// Mitsubishi GX Works2 project: 70常温静置库1130   PLC: Q10UDEH

TYPE BatteryCode : STRUCT
  arrwCode : ARRAY [0..8] OF WORD;
END_STRUCT END_TYPE

TYPE CommunicationIO : STRUCT
  i_iResponsPCPLC : INT;  (* 上位机写入-请求确认 *)
  i_iReadWriteFlagPCPLC : INT;  (* 上位机写入-读写标志位 *)
  i_iTaskProcessFlagPCPLC : INT;  (* 上位机写入-任务处理标志位 *)
  i_iCommandPCPLC : INT;  (* 上位机写入-命令字 *)
  i_iTaskIDPCPLC : INT;  (* 上位机写入-任务号 *)
  i_diDestinationDevicePCPLC : DINT;  (* 上位机写入-目标设备号 *)
  i_iProductIDPCPLC : INT;  (* 上位机写入-框码后4位 *)
  o_iRequestPLCPC : INT;  (* 上位机读取-请求状态 *)
  o_iReadWriteFlagPLCPC : INT;  (* 上位机读取-读写标志位 *)
  o_iDeviceStatusPLCPC : INT;  (* 上位机读取-设备状态 *)
  o_iTaskIDPLCPC : INT;  (* 上位机读取-任务号 *)
  o_iProductIDPLCPC : INT;  (* 上位机读取-框码后4位 *)
  i_iTypeInfoPCPLC : INT;  (* 上位机写入-批次标识，是否同批次 *)
  o_iForceInportPLCPC : INT;  (* 上位机读取-强制入库 *)
  o_iEmptyPLCPC : INT;  (* 上位机读取-有料状态 *)
  o_iFolderNumberPLCPC : INT;  (* 上位机读取-叠盘数量 *)
  i_xExtraCondition : BOOL;  (* 发送请求时的额外条件,比如需要升降到位 *)
  i_xExportConveyor : BOOL;  (* 线体是出库线体还是入库线体 *)
END_STRUCT END_TYPE

TYPE ConveyorIO : STRUCT
  xUnloadCCW : BOOL;  (* 下料为反转 *)
  xUnloadAlarm : BOOL;  (* 下料报警 *)
  xUnload : BOOL;  (* 下料请求 *)
  xPutInto : BOOL;  (* 线体直接投入物料 *)
  xNotArriveAlarm : BOOL;  (* 未到达报警 *)
  xNextRun : BOOL;  (* 下段线体运行 *)
  xMotorCW : BOOL;  (* 电机正转 *)
  xMotorCCW : BOOL;  (* 电机反转 *)
  xManual : BOOL;  (* 手动 *)
  xloadCCW : BOOL;  (* 上料为反转 *)
  xLimitAlarrm : BOOL;  (* 限位报警 *)
  xLoad : BOOL;  (* 上料请求 *)
  xForward : BOOL;  (* 正转手动 *)
  xEmpty : BOOL;  (* 线体状态为空 *)
  xCWPresent : BOOL;  (* 正转检测有无传感器 *)
  xCCWPresent : BOOL;  (* 反转检测有无传感器 *)
  xBusy : BOOL;  (* 工作中 *)
  xBackward : BOOL;  (* 反转手动 *)
  xAuto : BOOL;  (* 自动 *)
  xPosLimit : BOOL;  (* 正限位 *)
  xNegLimit : BOOL;  (* 负限位 *)
  xOverWidthAlarm : BOOL;  (* 超宽报警 *)
  xError : BOOL;  (* 报警 *)
  iProductCategoryIn : INT;  (* 产品类型输入 *)
  iProductCategory : INT;  (* 产品类型记录 *)
  iProductCategoryOut : INT;  (* 产品类型输出 *)
  diDeviceID : DINT;  (* 设备编号 *)
  tUnloadAlarmDelay : TIME;  (* 下料报警时间设置 *)
  tLoadDelay : TIME;  (* 上料延时设置 *)
  xSizeDeficientDetect : BOOL;  (* 尺寸缺陷检测 *)
  xZoneClear : BOOL;  (* 初始化线体清除 *)
  tZoneClearTime : TIME;  (* 初始化线体清除时间 *)
  iTaskIDIn : INT;  (* 产品类型输入 *)
  iTaskID : INT;  (* 产品类型记录 *)
  iTaskIDOut : INT;  (* 产品类型输出 *)
  diDesConveyorIn : DINT;  (* 产品类型输入 *)
  diDesConveyor : DINT;  (* 产品类型记录 *)
  diDesConveyorOut : DINT;  (* 产品类型输出 *)
END_STRUCT END_TYPE

TYPE FanucRobotIO : STRUCT
  o_xColumn : ARRAY [0..3] OF BOOL;  (* 行号 *)
  o_xRow : ARRAY [0..3] OF BOOL;  (* 列号 *)
  o_xPutNumber : ARRAY [0..3] OF BOOL;  (* 放料位 *)
  o_xSortStart : BOOL;  (* 开始启动 *)
  i_xPutOver : BOOL;  (* 放货完成 *)
  i_xPickOver : BOOL;  (* 取货完成 *)
  o_xCatchCylinder : BOOL;  (* 夹紧气缸 *)
  i_xBatteryDetect : ARRAY [0..3] OF BOOL;  (* 电池检测 *)
  i_xProtect : ARRAY [0..3] OF BOOL;  (* 限位保护 *)
END_STRUCT END_TYPE

TYPE FolderIO : STRUCT
  o_xCylinderGrabExtend : BOOL;  (* 气缸夹紧 *)
  o_xCylinderGrabRetract : BOOL;  (* 气缸松开 *)
  i_xCylinderGrabExtendDetect : BOOL;  (* 夹紧检测 *)
  i_xCylinderGrabRetractDetect : BOOL;  (* 松开检测 *)
  o_xCylinderUpExtend : BOOL;  (* 上层伸出 *)
  o_xCylinderUpRetract : BOOL;  (* 上层缩回 *)
  i_xCylinderUpExtendDetect : BOOL;  (* 上层伸出检测 *)
  i_xCylinderUpRetractDetect : BOOL;  (* 上层缩回检测 *)
  o_xCylinderDownExtend : BOOL;  (* 下层伸出 *)
  o_xCylinderDownRetract : BOOL;  (* 下层缩回 *)
  i_xCylinderDownExtendDetect : BOOL;  (* 下层伸出检测 *)
  i_xCylinderDownRetractDetect : BOOL;  (* 下层缩回检测 *)
  i_xExitEnable : BOOL;  (* 下料信号 *)
  i_xEntryEnable : BOOL;  (* 上料信号 *)
  o_xEntryPermit : BOOL;  (* 允许上料(拆盘需要，叠盘不需要) *)
  i_iFloor : INT;  (* 层数 *)
  i_xCylinderGrabExtendButton : BOOL;  (* 气缸夹紧按钮 *)
  i_xCylinderGrabRetractButton : BOOL;  (* 气缸松开按钮 *)
  i_xCylinderUpExtendButton : BOOL;  (* 上层伸出按钮 *)
  i_xCylinderUpRetractButton : BOOL;  (* 上层缩回按钮 *)
  i_xCylinderDownExtendButton : BOOL;  (* 下层伸出按钮 *)
  i_xCylinderDownRetractButton : BOOL;  (* 下层缩回按钮 *)
  o_xDownCylinderError : BOOL;  (* 下层气缸层伸出未到达 *)
  o_xUpCylinderError : BOOL;  (* 上层气缸伸出未到达 *)
  o_xGrabCylinderError : BOOL;  (* 夹紧气缸伸出未到达 *)
  i_tSetOvertime : TIME;  (* 未到达计时 *)
  o_xExitPremit : BOOL;  (* 允许下料(叠盘完成后输出) *)
  i_xTrayDetect : BOOL;  (* 托盘数量检测 *)
  i_NextConveyorEmpty : BOOL;  (* 下段线体空 *)
  i_FrontConveyorNextRun : BOOL;  (* 前段线体下料信号 *)
  m_iStepInput : INT;  (* 外部步骤输入 *)
  m_CountInput : INT;  (* 外部盘数量输入，只能输入0-3 *)
  o_CountResponsPC : INT;  (* 给上位机叠盘数量 *)
  i_FrontConveyorTypeInfo : INT;  (* 叠盘前扫码工位批次判断 *)
  o_RequestPC : INT;  (* 给上位机扫码请求 *)
  i_xFolderEnable : BOOL;  (* 叠盘使能，等于1时开始叠盘 *)
END_STRUCT END_TYPE

TYPE PackCommunicationIO : STRUCT
  i_iResponsPCPLC : INT;  (* 上位机写入-请求确认 *)
  i_iPackDoneAknPCPLC : INT;  (* 上位机写入-放行 *)
  i_iSinglePackResponsePCPLC : INT;  (* 上位机写入-单次装载应答 *)
  i_iSinglePackDoneAknPCPLC : INT;  (* 上位机写入-单次装载处理完成 *)
  o_iRequestPLCPC : INT;  (* 上位机读取-装载请求 *)
  o_iPackDonePLCPC : INT;  (* 上位机读取-装载完成 *)
  o_iSinglePackRequestPLCPC : INT;  (* 上位机读取-单次装载请求 *)
  o_iSinglePackDonePLCPC : INT;  (* 上位机读取-单次装载完成 *)
  o_iXCoordinatePLCPC : INT;  (* 上位机读取-行坐标 *)
  o_iYCoordinatePLCPC : INT;  (* 上位机读取-列坐标 *)
  o_arrwCode : ARRAY [0..7] OF BOOL;  (* 上位机读取-电芯码 *)
END_STRUCT END_TYPE

TYPE QueueElement : STRUCT
  xCondition : BOOL;
  iPriority : INT;
END_STRUCT END_TYPE

TYPE ShuttleCarIO : STRUCT
  xReady : BOOL;  (* 准备就绪 *)
  xForward : BOOL;  (* 正转 *)
  xBackward : BOOL;  (* 反转 *)
  iCurrentPos : INT;  (* 当前位置 *)
  iDestinationPos : INT;  (* 目标位置 *)
  xCW : BOOL;  (* 正转输出 *)
  xCCW : BOOL;  (* 反转输出 *)
  xBrake : BOOL;  (* 刹车 *)
  xHomeSwitch : BOOL;  (* 零位接近开关 *)
  xPosLimit : BOOL;  (* 正限位 *)
  xNegLimit : BOOL;  (* 负限位 *)
  xMDIExe : BOOL;  (* MDI开始 *)
  xMDIDone : BOOL;  (* MDI 完成 *)
  xPassLimit : BOOL;  (* 限位屏蔽 *)
  xPosLimitCatch : BOOL;  (* 正限位捕捉 *)
  xNegLimitCatch : BOOL;  (* 负限位捕捉 *)
  xHomeExe : BOOL;  (* 开始寻零 *)
  xHomeDone : BOOL;  (* 寻零完成 *)
  xHomeBusy : BOOL;  (* 寻零中 *)
  xHomeFailed : BOOL;  (* 寻零失败 *)
  xBusy : BOOL;  (* 工作中 *)
  tArriveDelay : TIME;  (* 到位延时 *)
  xCylinder : BOOL;  (* 气缸控制 *)
  tBrakeDelay : TIME;  (* 抱闸延时 *)
  xPauseRamp : BOOL;  (* 暂停减速斜坡标志位 *)
  xPresentDetect1 : BOOL;  (* 物料有无检测1 *)
  xPresentDetect2 : BOOL;  (* 物料有无检测2 *)
  xOvertimeAlarm : BOOL;  (* 超时报警 *)
  tSetOverTime : TIME;  (* 设置超时时间 *)
  xLooseDetect : BOOL;  (* 松绳检测 *)
  xLooseAlarm : BOOL;  (* 松绳报警 *)
  xArrive : BOOL;  (* 到位信号 *)
  diDeviceID : DINT;  (* 设备编号 *)
  xMoveStep : BOOL;  (* 寸动 *)
  xAdrSwitch : ARRAY [1..8] OF BOOL;  (* 位置开关 *)
END_STRUCT END_TYPE

TYPE SortCommunicationIO : STRUCT
  i_iResponsPCPLC : INT;  (* 上位机写入-应答 *)
  i_iSortDoneAknPCPLC : INT;  (* 上位机写入-任务处理完成 *)
  i_arriBatteryStatus : ARRAY [1..128] OF INT;  (* 上位机写入-电池状态 *)
  o_iRequestPLCPC : INT;  (* 上位机读取-请求 *)
  o_iSortDonePLCPC : INT;  (* 上位机读取-分拣完成 *)
  i_iInfoWriteDone : INT;  (* 上位机写入-参数写入完成 *)
  i_xSortOver : BOOL;  (* 按钮，分拣完成 *)
  o_xSortDone : BOOL;  (* 状态，分拣完成 *)
END_STRUCT END_TYPE

TYPE SwitchIO : STRUCT
  xLiftCylinderRetractDetect : BOOL;
  xLiftCylinderExtendDetect : BOOL;
  xLiftCylinderRetract : BOOL;
  xLiftCylinderExtend : BOOL;
  xEntryBarCylinderRetract : BOOL;
  xLiftCylinderExtendInit : BOOL;
  xEntryEnable : BOOL;
  xExitEnable : BOOL;
  xExitBarCylinderRetract : BOOL;
  xSwithEnable : BOOL;
  xLiftCylinderRetractButton : BOOL;
  xLiftCylinderExtendButton : BOOL;
  xEntryBarCylinderRetractButton : BOOL;
  xExitBarCylinderRetractButton : BOOL;
  xPutInto : BOOL;  (* 单体复位 *)
  tSetOvertime : TIME;  (* 设定超时报警时间 *)
  xOvertimeAlarm : BOOL;  (* 超时报警 *)
END_STRUCT END_TYPE

TYPE UConveyorIO : STRUCT
  xLiftCylinderRetractDetect1 : BOOL;
  xLiftCylinderRetractDetect2 : BOOL;
  xLiftCylinderExtendDetect1 : BOOL;
  xLiftCylinderExtendDetect2 : BOOL;
  xLiftCylinderRetract1 : BOOL;
  xLiftCylinderRetract2 : BOOL;
  xLiftCylinderExtend1 : BOOL;
  xLiftCylinderExtend2 : BOOL;
  xExitBarCylinderRetract1 : BOOL;
  xExitBarCylinderRetract2 : BOOL;
  xLiftCylinderExtendInit1 : BOOL;
  xLiftCylinderExtendInit2 : BOOL;
  xEntryEnable1 : BOOL;
  xEntryEnable2 : BOOL;
  xEntryEnable3 : BOOL;
  xExitEnable1 : BOOL;
  xExitEnable2 : BOOL;
  xExitEnable3 : BOOL;
  xPassEnable : BOOL;  (* 直接放行去下段 *)
  xLiftCylinderRetractButton1 : BOOL;
  xLiftCylinderRetractButton2 : BOOL;
  xLiftCylinderExtendButton1 : BOOL;
  xLiftCylinderExtendButton2 : BOOL;
  xExitBarCylinderRetractButton1 : BOOL;
  xExitBarCylinderRetractButton2 : BOOL;
  xPutInto : BOOL;  (* 单体复位 *)
  tSetOvertime : TIME;  (* 设定超时报警时间 *)
  xOvertimeAlarm : BOOL;  (* 超时报警 *)
  iTask : INT;  (* 3个任务 *)
  xBatteryDetect1 : BOOL;  (* 电池检测1 *)
  xBatteryDetect2 : BOOL;  (* 电池检测2 *)
  xBatteryError : BOOL;  (* 空框里有电池错误 *)
END_STRUCT END_TYPE

TYPE ServoIO : STRUCT
  xQD75Ready : BOOL;  (* QD75Ready---X0 *)
  xQD75Error1 : BOOL;  (* 1轴出错---X8 *)
  xQD75Error2 : BOOL;  (* 2轴出错---X9 *)
  xQD75Error3 : BOOL;  (* 3轴出错---XA *)
  xQD75Error4 : BOOL;  (* 4轴出错---XB *)
  xQD75Busy1 : BOOL;  (* 1轴BUSY---XC *)
  xQD75Busy2 : BOOL;  (* 2轴BUSY---XD *)
  xQD75Busy3 : BOOL;  (* 3轴BUSY---XE *)
  xQD75Busy4 : BOOL;  (* 4轴BUSY---XF *)
  xQD75Starting1 : BOOL;  (* 1轴起动完成---X10 *)
  xQD75Starting2 : BOOL;  (* 2轴起动完成---X11 *)
  xQD75Starting3 : BOOL;  (* 3轴起动完成---X12 *)
  xQD75Starting4 : BOOL;  (* 4轴起动完成---X13 *)
  xQD75LocateDone1 : BOOL;  (* 1轴定位完成---X14 *)
  xQD75LocateDone2 : BOOL;  (* 2轴定位完成---X15 *)
  xQD75LocateDone3 : BOOL;  (* 3轴定位完成---X16 *)
  xQD75LocateDone4 : BOOL;  (* 4轴定位完成---X17 *)
  xQD75Stop1 : BOOL;  (* 1轴停止---Y4 *)
  xQD75Stop2 : BOOL;  (* 2轴停止---Y5 *)
  xQD75Stop3 : BOOL;  (* 3轴停止---Y6 *)
  xQD75Stop4 : BOOL;  (* 4轴停止---Y7 *)
  xQD75JogCW1 : BOOL;  (* 1轴JOG正转---Y8 *)
  xQD75JogCCW1 : BOOL;  (* 1轴JOG反转---Y9 *)
  xQD75JogCW2 : BOOL;  (* 2轴JOG正转---YA *)
  xQD75JogCCW2 : BOOL;  (* 2轴JOG反转---YB *)
  xQD75JogCW3 : BOOL;  (* 3轴JOG正转---YC *)
  xQD75JogCCW3 : BOOL;  (* 3轴JOG反转---YD *)
  xQD75JogCW4 : BOOL;  (* 4轴JOG正转---YE *)
  xQD75JogCCW4 : BOOL;  (* 4轴JOG反转---YF *)
  xQD75LocateStart1 : BOOL;  (* 1轴定位起动---Y10 *)
  xQD75LocateStart2 : BOOL;  (* 2轴定位起动---Y11 *)
  xQD75LocateStart3 : BOOL;  (* 3轴定位起动---Y12 *)
  xQD75LocateStart4 : BOOL;  (* 4轴定位起动---Y13 *)
  xQD75Ban1 : BOOL;  (* 1轴禁止---Y14 *)
  xQD75Ban2 : BOOL;  (* 2轴禁止---Y15 *)
  xQD75Ban3 : BOOL;  (* 3轴禁止---Y16 *)
  xQD75Ban4 : BOOL;  (* 4轴禁止---Y17 *)
  diQD75CurrentPos1 : DINT;  (* 1轴当前位置(QD75-PLC)---U0\G800 *)
  diQD75LastPos1 : DINT;  (* 1轴1S前的位置，方便确认是否有输出 *)
  iQD75ErrorNumber1 : INT;  (* 1轴错误代码(QD75-PLC)---U0\G806 *)
  iQD75AlarmNumber1 : INT;  (* 1轴警告代码(QD75-PLC)---U0\G807 *)
  iQD75State1 : INT;  (* 1轴运行状态(QD75-PLC)---U0\G809 *)
  diQD75Speed1 : DINT;  (* 1轴速度(QD75-PLC)---U0\G810 *)
  diQD75DestinationPos1 : DINT;  (* 1轴目标地址(QD75-PLC)---U0\G818 *)
  iQD75DestiNumber1 : INT;  (* 1轴定位目标编号(QD75-PLC)---U0\G835 *)
  iQD75LastNumber1 : INT;  (* 1轴上次定位编号(QD75-PLC)---U0\G837 *)
  iLocateStartNumber1 : INT;  (* 1轴定位起动编号(PLC-QD75)---U0\G1500 *)
  iReset1 : INT;  (* 1轴出错给1复位(PLC-QD75)---U0\G1502 *)
  iReStart1 : INT;  (* 1轴给1重起动(PLC-QD75)---U0\G1503 *)
  diJOGSpeed1 : DINT;  (* 1轴JOG速度(PLC-QD75)---U0\G1518 *)
  xPLCReady : BOOL;  (* PLCReady--Y0 *)
  diQD75CurrentPos3 : DINT;  (* 3轴当前位置(QD75-PLC)---U0\G1000 *)
  diQD75LastPos3 : DINT;  (* 3轴1S前的位置，方便确认是否有输出 *)
  iQD75ErrorNumber3 : INT;  (* 3轴错误代码(QD75-PLC)---U0\G1006 *)
  iQD75AlarmNumber3 : INT;  (* 3轴警告代码(QD75-PLC)---U0\G1007 *)
  iQD75State3 : INT;  (* 3轴运行状态(QD75-PLC)---U0\G1009 *)
  diQD75Speed3 : DINT;  (* 3轴速度(QD75-PLC)---U0\G1010 *)
  diQD75DestinationPos3 : DINT;  (* 3轴目标地址(QD75-PLC)---U0\G1018 *)
  iQD75DestiNumber3 : INT;  (* 3轴定位目标编号(QD75-PLC)---U0\G1035 *)
  iQD75LastNumber3 : INT;  (* 3轴上次定位编号(QD75-PLC)---U0\G1037 *)
  iLocateStartNumber3 : INT;  (* 3轴定位起动编号(PLC-QD75)---U0\G1700 *)
  iReset3 : INT;  (* 3轴出错给1复位(PLC-QD75)---U0\G1702 *)
  iReStart3 : INT;  (* 3轴给1重起动(PLC-QD75)---U0\G1703 *)
  diJOGSpeed3 : DINT;  (* 3轴JOG速度(PLC-QD75)---U0\G1718 *)
  diQD75CurrentPos2 : DINT;  (* 2轴当前位置(QD75-PLC)---U0\G900 *)
  diQD75LastPos2 : DINT;  (* 2轴1S前的位置，方便确认是否有输出 *)
  iQD75ErrorNumber2 : INT;  (* 2轴错误代码(QD75-PLC)---U0\G906 *)
  iQD75AlarmNumber2 : INT;  (* 2轴警告代码(QD75-PLC)---U0\G907 *)
  iQD75State2 : INT;  (* 2轴运行状态(QD75-PLC)---U0\G909 *)
  diQD75Speed2 : DINT;  (* 2轴速度(QD75-PLC)---U0\G910 *)
  diQD75DestinationPos2 : DINT;  (* 2轴目标地址(QD75-PLC)---U0\G918 *)
  iQD75DestiNumber2 : INT;  (* 2轴定位目标编号(QD75-PLC)---U0\G935 *)
  iQD75LastNumber2 : INT;  (* 2轴上次定位编号(QD75-PLC)---U0\G937 *)
  iLocateStartNumber2 : INT;  (* 2轴定位起动编号(PLC-QD75)---U0\G1600 *)
  iReset2 : INT;  (* 2轴出错给1复位(PLC-QD75)---U0\G1602 *)
  iReStart2 : INT;  (* 2轴给1重起动(PLC-QD75)---U0\G1603 *)
  diJOGSpeed2 : DINT;  (* 2轴JOG速度(PLC-QD75)---U0\G1618 *)
  diQD75CurrentPos4 : DINT;  (* 4轴当前位置(QD75-PLC)---U0\G1100 *)
  diQD75LastPos4 : DINT;  (* 4轴1S前的位置，方便确认是否有输出 *)
  iQD75ErrorNumber4 : INT;  (* 4轴错误代码(QD75-PLC)---U0\G1106 *)
  iQD75AlarmNumber4 : INT;  (* 4轴警告代码(QD75-PLC)---U0\G1107 *)
  iQD75State4 : INT;  (* 4轴运行状态(QD75-PLC)---U0\G1109 *)
  diQD75Speed4 : DINT;  (* 4轴速度(QD75-PLC)---U0\G1110 *)
  diQD75DestinationPos4 : DINT;  (* 4轴目标地址(QD75-PLC)---U0\G1118 *)
  iQD75DestiNumber4 : INT;  (* 4轴定位目标编号(QD75-PLC)---U0\G1135 *)
  iQD75LastNumber4 : INT;  (* 4轴上次定位编号(QD75-PLC)---U0\G1137 *)
  iLocateStartNumber4 : INT;  (* 4轴定位起动编号(PLC-QD75)---U0\G1800 *)
  iReset4 : INT;  (* 4轴出错给1复位(PLC-QD75)---U0\G1802 *)
  iReStart4 : INT;  (* 4轴给1重起动(PLC-QD75)---U0\G1803 *)
  diJOGSpeed4 : DINT;  (* 4轴JOG速度(PLC-QD75)---U0\G1818 *)
  xResetServo : BOOL;  (* 重新启动 *)
  xBackHome1 : BOOL;  (* 1轴回原点信号 *)
  xBackHome2 : BOOL;  (* 2轴回原点信号 *)
  xBackHome3 : BOOL;  (* 3轴回原点信号 *)
  xBackHome4 : BOOL;  (* 4轴回原点信号 *)
END_STRUCT END_TYPE

// global labels: Global
VAR_GLOBAL
  g_xAuto AT M11 : BOOL;
  g_xManual : BOOL;
  g_xEStop AT X0 : BOOL;
  g_xReset AT X3 : BOOL;
  g_xStackLampRed AT Y200 : BOOL;
  g_xStackLampAmber AT Y201 : BOOL;
  g_xStackLampGreen AT Y202 : BOOL;
  g_xBuzzer AT Y203 : BOOL;
  g_xStop AT X3 : BOOL;
  g_xAutoStart AT X2 : BOOL;
  g_xRemoteAutoStart AT M0 : BOOL;
  g_xRemoteAuto AT M10 : BOOL;
  g_iState AT D40 : INT;
  g_iLocalAutoStep : BOOL;
  g_xAlarm : BOOL;
  g_xPause AT M3 : BOOL;  (* 暂停 *)
  g_diDeviceIDSelect AT D0 : DINT;
  g_xResetSingle AT M4 : BOOL;  (* 单线体复位 *)
  g_xInsertTask AT M5 : BOOL;  (* 插入任务 *)
  g_iInsertTaskID AT D2 : INT;  (* 插入任务号 *)
  g_iConveyorStatus AT D4 : INT;
  g_iInsertCategory AT D6 : INT;
  g_diInsertDesConveyor AT D8 : DINT;
  g_xRGVTcpFailed : BOOL;
  g_xAutoLamp AT Y204 : BOOL;
  g_xAutoSwitch AT X1 : BOOL;
  g_xMute : BOOL;
  g_xResetTask1 AT M9 : BOOL;  (* 复位排队任务的 *)
  g_x60TcpFailed : BOOL;
  m_Ocv2_1Forbidden AT M990 : BOOL;  (* OCV2-1禁用 *)
  m_Ocv2_2Forbidden AT M991 : BOOL;  (* OCV2-2禁用 *)
  m_Choose1Forbidden AT M992 : BOOL;  (* 挑选1禁用 *)
  m_Ocv3_1Forbidden AT M993 : BOOL;  (* OCV3-1禁用 *)
  m_Ocv3_2Forbidden AT M994 : BOOL;  (* OCV3-2禁用 *)
  m_Choose2Forbidden AT M995 : BOOL;  (* 挑选2禁用 *)
  g_xRGVRemoteAuto AT M20 : BOOL;  (* RGV远程自动 *)
  g_SemiStart AT M21 : BOOL;
END_VAR

// task Task1 (event TRUE, interval 0, priority 31): POU, START, TCP

FUNCTION_BLOCK Conveyor
VAR
  m_xPresentDelay : BOOL;  (* 有无判断延时 *)
  m_xLoadDelayOut : BOOL;  (* 上料延时输出 *)
  m_xInitial : BOOL;  (* 初始化 *)
  m_tUnloadTimer : TIME;  (* 下料计时器 *)
  m_tPresentDelayCurrentTime : TIME;
  m_tonUnloadAlam : TON;  (* 下料报警定时器 *)
  m_tonPresentDelay : TON;  (* 物料有无判断延时，防止误动作 *)
  m_tonNotArriveAlarm : TON;  (* 未到达报警计时 *)
  m_tonLoadDelay : TON;  (* 上料延时 *)
  m_tNotArriveCurrentTime : TIME;  (* 未到达报警计时当前时间 *)
  m_tLoadTimer : TIME;  (* 上料计时器 *)
  iStep : INT;  (* 上料步骤 *)
  m_wStateWord : INT;
END_VAR
VAR_IN_OUT
  ConveyorMotor : ConveyorIO;  (* 输送线输入输出 *)
END_VAR
VAR
  m_tonZoneClear : TON;  (* 初始化清除 *)
  m_tZoneClearCurrentTime : TIME;  (* 初始化清除当前时间 *)
  m_xAutoClear : BOOL;  (* 初始化清除标志位 *)
  m_xZoneClearDone : BOOL;  (* 初始化清除完成 *)
END_VAR
(*////////////////////////////////////////////////////////////////////////////////////////////////////////////
//传输线控制FB块，可控制单方向线体，双向旋转线体，支持双向上下料            
//线体初始化后为空的情况下输入xLoad信号即可进行上料动作，使用xLoadCCW信号可反方向上料
//增加了产品信息和产品种类的储存，当传输线为空和上料进行标志位为零的情况下清除产品信息和产品种类
//使用方式是在置位xLoad信号后，把产品信息和产品种类传入，等下料后自动清零
//线体不为空的情况下使用xUnload信号可进行下料动作，物料有无传感器的下降沿后出发计时器，延时断开传输线旋转
//单方向传输线体把xLoadCCW、xUnloadCCW设置为零，双向线体上料方向和下料反向的,方向固定的 把xUnloadCCW设置为1
//双方向线体双向都能上下料的要根据上料的方向来设置xLoadCCW,xUnloadCCW
//增加工作中信号xBusy当电机正转 显示为工作中
//增加上下料超时报警，xLoadAlarm，xUnloadAlarm，设定时间在LOAD_UNLOAD_TIME常量上，现在设置的为30秒
//增加xPutInto信号，用于直接投入的物料，检测开关感应到后，直接进入下料流程，上升沿有效
//离开延时改为变量 iLeaveDelay 默认为0 离开检测开关离输送线尾端比较远的线体需要根据情况设定100ms为单位
//增加初始化标志位，增加进入延时时间，初始化为进入延时时间为0 ，离开延时时间为2S，通过外围接口可以更改
//修改信息  修改后请增加版本
//12-17进行了优化，增加了未到达报警，当物料未传送到下一设备，就报未到达报警，使用xNextRun标志位制作，没有正常到达
//第0步，不能跳转到第一步把标志位复位，即出现中断情况，2秒后报警
//修改信息  修改后请增加版本
//上料延时增加为50ms防止干扰信号
//nextrun信号在 第三步也要复位
//增加限位报警
//增加超宽报警
//增加产品型号输出在下料的时候把产品型号输送给下一段线体
//增加线体单独复位
//增加任务插入功能配合全局变量
//增加暂停功能
//增加线体状态字显示  0 空闲 1：有料  2 工作中  3  超限报警 4 超宽报警  5 未到达报警  6 下料超时报警
//空料判断放在自动前，进行有无报警判断，然后跳转
//修改超限报警，与尺寸检测报警
////YAO      V1.0
//把所有的IF语句去掉，  IF语句占用指针存储区，容易造成存储区不足的现象
////YAO      V1.1
//初始化清除线体标志位xZoneClear
//ZPA zero pressure accumulation  Term that describes the Conveyor controls and mechanical scheme that will 
//cause loads to queue on a conveyor in discrete zones such that loads do not touch each other(wrapped boxed tray tote carton)
//除了产品信息外，还增加了目标地址，任务类型的数据传递。
//YAO      V1.0
///////////////////////////////////////////////////////////////////////////////////////////////////////////
(*********************************************************)
(*//初始化，
//上料延时位0S，下料报警延时为30S
//下料延时设一个比较大的时间，主要依靠xunload标志位来停止输送线，特殊情况可以用延时来停止物流线下料
//设置时间大的时候计时器会失效*)
IF NOT m_xInitial THEN
	ConveyorMotor.tLoadDelay:=T#100ms;
	ConveyorMotor.tUnloadAlarmDelay:=T#30s;
	ConveyorMotor.xPosLimit:=1;
	ConveyorMotor.xNegLimit:=1;
	ConveyorMotor.xSizeDeficientDetect:=0;
	ConveyorMotor.xZoneClear:=0;
	ConveyorMotor.tZoneClearTime:=T#10s;
	m_xInitial:=1;
END_IF;
(*//自动
//复位信号把步号置0，但xLoad与xUnload没有复位，调用程序需要注意复位后把这两个信号置零，以免发生误动作
//物料有无判断增加延时，防止开自动瞬间误动作发生*)
m_tonPresentDelay(IN:= ConveyorMotor.xCWPresent OR ConveyorMotor.xCCWPresent,
 PT:=T#100ms,
 Q:= m_xPresentDelay,
 ET:= m_tPresentDelayCurrentTime);
CASE iStep OF
0:(*//初始化*)
	ConveyorMotor.xMotorCW:=0;
	ConveyorMotor.xMotorCCW:=0;
	ConveyorMotor.xNextRun:=0;
	ConveyorMotor.iProductCategoryOut:=0;
	ConveyorMotor.iTaskIDOut:=0;
	ConveyorMotor.diDesConveyorOut:=0;
	out(NOT m_xPresentDelay,ConveyorMotor.xEmpty);(*	//判断物料有无传感器*)	
	mov(m_xPresentDelay AND g_xAuto AND NOT ConveyorMotor.xError,3,iStep);(*//自动情况下进行跳转*)(*无超限报警*)
	mov(NOT m_xPresentDelay AND g_xAuto AND NOT ConveyorMotor.xError,1,iStep);
1: (*//上料*)
	rst(ConveyorMotor.xLoad ,ConveyorMotor.iProductCategory);(*//上料开始清除产品信息*)
	rst(ConveyorMotor.xLoad ,ConveyorMotor.iTaskID);
	rst(ConveyorMotor.xLoad ,ConveyorMotor.diDesConveyor);
	mov(ConveyorMotor.xLoad,2,iStep);
2: (*//上料完成*)
	ConveyorMotor.iProductCategory:=ConveyorMotor.iProductCategoryIn;(* //产品信息传入*)
	ConveyorMotor.iTaskID:=ConveyorMotor.iTaskIDIn;
	ConveyorMotor.diDesConveyor:=ConveyorMotor.diDesConveyorIn;
	set(ConveyorMotor.xloadCCW,ConveyorMotor.xMotorCCW);
	rst(ConveyorMotor.xloadCCW,ConveyorMotor.xMotorCW);
	set(NOT ConveyorMotor.xloadCCW,ConveyorMotor.xMotorCW);
	rst(NOT ConveyorMotor.xloadCCW,ConveyorMotor.xMotorCCW);	
	m_tonLoadDelay(IN:= (ConveyorMotor.xCWPresent AND NOT ConveyorMotor.xloadCCW) 
  		OR (ConveyorMotor.xCCWPresent AND ConveyorMotor.xloadCCW) ,
  PT:= ConveyorMotor.tLoadDelay ,
  Q:= m_xLoadDelayOut ,
  ET:= m_tLoadTimer );
	mov(m_xLoadDelayOut,3, iStep);
3:(*//下料请求*)	
	ConveyorMotor.xMotorCW:=0;
	ConveyorMotor.xMotorCCW:=0;
	ConveyorMotor.xEmpty:=0;
	mov(ConveyorMotor.xUnload AND NOT ConveyorMotor.xOverWidthAlarm,4,iStep);
4:(*	//下料完成*)
	set(ConveyorMotor.xUnloadCCW,ConveyorMotor.xMotorCCW);
	rst(ConveyorMotor.xUnloadCCW,ConveyorMotor.xMotorCW);
	set(NOT ConveyorMotor.xUnloadCCW,ConveyorMotor.xMotorCW);
	rst(NOT ConveyorMotor.xUnloadCCW,ConveyorMotor.xMotorCCW);	
	ConveyorMotor.xNextRun:=1; (*下一段线体旋转*)
	ConveyorMotor.iProductCategoryOut:=ConveyorMotor.iProductCategory;(*产品型号输出给下一段线体*)
	ConveyorMotor.iTaskIDOut:=ConveyorMotor.iTaskID;
	ConveyorMotor.diDesConveyorOut:=ConveyorMotor.diDesConveyor;
	mov( NOT ConveyorMotor.xUnload , 0, istep );
END_CASE;
(*In-feed zone clear and ready to accept a load from upstream Conveyor*)
set(ldp(TRUE,g_xAuto) ,m_xAutoClear);
rst(ldf(TRUE,g_xAuto) ,m_xAutoClear);
m_tonZoneClear(IN:= m_xAutoClear AND ConveyorMotor.xZoneClear ,PT:= ConveyorMotor.tZoneClearTime ,Q:=m_xZoneClearDone ,ET:= m_tZoneClearCurrentTime );
set(m_xAutoClear AND ConveyorMotor.xZoneClear,ConveyorMotor.xMotorCW);
mov( m_xAutoClear AND ConveyorMotor.xZoneClear, 0 ,iStep );
rst(  ldf(TRUE, m_xAutoClear ) ,ConveyorMotor.xMotorCW);
rst( m_xZoneClearDone OR m_xPresentDelay  , m_xAutoClear );
(*投入上料，搬出下料，也可用来初始化*)
movp( ConveyorMotor.xPutInto, 0 , iStep );
(*//当前任务显示*)
movp( ConveyorMotor.diDeviceID=g_diDeviceIDSelect , ConveyorMotor.iProductCategory , g_iInsertCategory );
movp( ConveyorMotor.diDeviceID=g_diDeviceIDSelect , ConveyorMotor.iTaskID , g_iInsertTaskID );
dmovp( ConveyorMotor.diDeviceID=g_diDeviceIDSelect , ConveyorMotor.diDesConveyor , g_diInsertDesConveyor );
(*//插入任务*)
mov(g_xInsertTask AND ConveyorMotor.diDeviceID=g_diDeviceIDSelect ,g_iInsertCategory , ConveyorMotor.iProductCategory );
mov(g_xInsertTask AND ConveyorMotor.diDeviceID=g_diDeviceIDSelect , g_iInsertTaskID , ConveyorMotor.iTaskID );
dmov(g_xInsertTask AND ConveyorMotor.diDeviceID=g_diDeviceIDSelect , g_diInsertDesConveyor , ConveyorMotor.diDesConveyor );
(*//单线体复位，当设备号与本线体一致的时候执行复位*)
mov(g_xResetSingle AND ConveyorMotor.diDeviceID=g_diDeviceIDSelect , 0 , iStep );
rst(g_xResetSingle AND ConveyorMotor.diDeviceID=g_diDeviceIDSelect ,ConveyorMotor.xNextRun );
rst(g_xResetSingle AND ConveyorMotor.diDeviceID=g_diDeviceIDSelect  ,ConveyorMotor.xLimitAlarrm );
rst(g_xResetSingle AND ConveyorMotor.diDeviceID=g_diDeviceIDSelect  ,ConveyorMotor.xOverWidthAlarm );
(*//手动*)
(*//正转*)
set( g_xManual   
AND ConveyorMotor.xForward 
AND ConveyorMotor.xBackward=0 
AND ConveyorMotor.xMotorCCW=0 
AND g_xEStop  , 
ConveyorMotor.xMotorCW);
rst((g_xManual 
AND (NOT ConveyorMotor.xForward  
OR ConveyorMotor.xBackward 
OR ConveyorMotor.xMotorCCW )) 
OR  NOT g_xEStop,
ConveyorMotor.xMotorCW);
(*//反转*)		
set(g_xManual 
AND ConveyorMotor.xBackward 
AND ConveyorMotor.xForward=0 
AND ConveyorMotor.xMotorCW=0 
AND g_xEStop ,
ConveyorMotor.xMotorCCW);
rst((g_xManual AND 
(NOT ConveyorMotor.xBackward  
OR ConveyorMotor.xForward 
OR ConveyorMotor.xMotorCW ) ) 
OR NOT g_xEStop,
ConveyorMotor.xMotorCCW);
mov(g_xManual ,0,iStep);(*//手动后上下料程序步骤清零*)
(*暂停*)
rst(g_xPause,ConveyorMotor.xMotorCCW);
rst( g_xPause , ConveyorMotor.xMotorCW );
(*工作中信号输出*)
ConveyorMotor.xBusy:=ConveyorMotor.xMotorCCW OR ConveyorMotor.xMotorCW;
(*//未到达报警*)
m_tonNotArriveAlarm(IN:= iStep=0 AND ConveyorMotor.xNextRun  ,PT:= T#2s,Q:= ConveyorMotor.xNotArriveAlarm ,ET:= m_tNotArriveCurrentTime );
(*//下料超时报警*)
m_tonUnloadAlam(IN:= iStep=4,PT:=ConveyorMotor.tUnloadAlarmDelay,Q:= ConveyorMotor.xUnloadAlarm,ET:=m_tUnloadTimer );
(*//限位报警,进料检测开关失效*)
set(  ( ((ConveyorMotor.xloadCCW AND NOT ConveyorMotor.xNegLimit)            (*反转上料，碰到负限位*)
			OR  ( NOT ConveyorMotor.xloadCCW AND NOT ConveyorMotor.xPosLimit)) (*正转上料，碰到正限位*)
		AND iStep=2) (*上料过程*)
	OR
	( iStep=4 (*下料过程*)
		AND( (ConveyorMotor.xUnloadCCW AND NOT ConveyorMotor.xPosLimit)  
			OR (NOT ConveyorMotor.xUnloadCCW AND NOT ConveyorMotor.xNegLimit)))  ,  
	ConveyorMotor.xLimitAlarrm );
mov( ( ((ConveyorMotor.xloadCCW AND NOT ConveyorMotor.xNegLimit)            (*反转上料，碰到负限位*)
			OR  ( NOT ConveyorMotor.xloadCCW AND NOT ConveyorMotor.xPosLimit)) (*正转上料，碰到正限位*)
		AND iStep=2) (*上料过程*)
	OR
	( iStep=4 (*下料过程*)
		AND( (ConveyorMotor.xUnloadCCW AND NOT ConveyorMotor.xPosLimit)  
			OR (NOT ConveyorMotor.xUnloadCCW AND NOT ConveyorMotor.xNegLimit)))  ,
	0,
	iStep);
(*//超宽报警*)
set( (iStep=3 OR iStep=1) AND (NOT ConveyorMotor.xNegLimit OR NOT ConveyorMotor.xPosLimit) , ConveyorMotor.xOverWidthAlarm  );
(*//尺寸不足报警*)
(*//有料状态下检测两个开关都要有信号*)
set( iStep=3 AND ConveyorMotor.xSizeDeficientDetect AND (NOT ConveyorMotor.xCCWPresent OR NOT ConveyorMotor.xCWPresent) ,  ConveyorMotor.xOverWidthAlarm );
mov( iStep=3 AND ConveyorMotor.xSizeDeficientDetect AND (NOT ConveyorMotor.xCCWPresent OR NOT ConveyorMotor.xCWPresent),0,iStep);
(*//总报警*)
ConveyorMotor.xError:=ConveyorMotor.xLimitAlarrm
 OR ConveyorMotor.xNotArriveAlarm
 OR ConveyorMotor.xUnloadAlarm                                             
 OR ConveyorMotor.xOverWidthAlarm;

(*//状态输出*)(*状态显示，容易造成指针容量不足*)
mov( ConveyorMotor.xEmpty AND NOT ConveyorMotor.xBusy , 0 , m_wStateWord);
mov( ConveyorMotor.xEmpty=0 ,  		1 , m_wStateWord);
mov( ConveyorMotor.xBusy ,  			2 , m_wStateWord);
mov( ConveyorMotor.xLimitAlarrm ,  	3, 	m_wStateWord);
mov(ConveyorMotor.xOverWidthAlarm ,  4 , m_wStateWord);
mov( ConveyorMotor.xNotArriveAlarm ,  5 , m_wStateWord);
mov( ConveyorMotor.xUnloadAlarm,  	6 , m_wStateWord);
(*选择本线体后，将状态赋值给全局变量进行显示*)
mov( ConveyorMotor.diDeviceID=g_diDeviceIDSelect , m_wStateWord, g_iConveyorStatus );
END_FUNCTION_BLOCK

FUNCTION_BLOCK ConveyorCommunication
VAR_IN_OUT
  ConveyorIO : ConveyorIO;
  CommunicationIO : CommunicationIO;
END_VAR
VAR_OUTPUT
  o_iErrorNub : INT;  (* 错误代码 *)
  o_xReqSuccess : BOOL;  (* 请求成功 *)
END_VAR
VAR
  m_xInitial : BOOL;  (* 初始化 *)
  o_xError : BOOL;  (* 通信数据错误 *)
END_VAR
(********************************************************************************)
(*
DB1区(PC->PLC)15个字		
"字(16位）序号
(从1开始)"			功能描述											具体参数解释
1					请求确认	"										1：复位
				 														2：读码(入库申请）成功
				 														3：取放货完成 
																		4：旋转
																		5：不旋转
																		101：条码空
																		102：条码规则校验失败
																		103：步号校验失败
																		104：无库位可用 
"
2	预留	
3	预留	
4	预留	
5	预留	
6	读写标志位	"														1：写入数据
																		2：读数据完成"
7	任务处理标志	"														１：复位
																		２：完成"
8	命令字	"
																		21-送出（任务起点与终点不同，即向下一台输送机移载）
																		22：叠盘
"
9	任务号	"															1~65535唯一任务标识"
10	目标设备号															只有送出任务才有效
11		
12	筐码后4位	
				

DB2区(PLC->PC)15个字			
"字(16位）序号
(从1开始)"	功能描述	具体参数解释	
1	请求状态	"１：复位
２：请求"	实时状态，没有时序交互
2	强制入库(预留）	"１：复位
２：强制入库"	
3	预留(叠盘数量）	只对叠盘工位有效	
4	预留		
5			
6	读写标志位	"1：写入数据
2：读数据完成"	"有交互
时序"
7	设备状态	"1:空闲
2：工作中
3:任务完成（只有目标设备才会报任务完成）
４：故障"	
8	任务号	1~65535唯一任务标识，当输送任务执行完成后，将PC下发的任务号上报	
9	筐码后4位		
10	预留		
11			
			





2018.8.3 YAO 1.0
*)
(********************************************************************************)
(*如果外部不设置，就认为没有额外条件，有料就请求*)
IF NOT m_xInitial THEN
		CommunicationIO.i_xExtraCondition:=1;
		CommunicationIO.i_xExportConveyor:=0;
		m_xInitial:=1;
END_IF;
(*//有料状态*)
IF ConveyorIO.xEmpty THEN
	CommunicationIO.o_iEmptyPLCPC:=1;
	CommunicationIO.o_iRequestPLCPC:=1;(*无料撤销请求*)
	ELSE
	CommunicationIO.o_iEmptyPLCPC:=2;
END_IF;

(*//请求状态*)
(*入库段线体*)
IF CommunicationIO.i_xExportConveyor=0 THEN
		IF NOT ConveyorIO.xEmpty AND CommunicationIO.i_xExtraCondition THEN
			CommunicationIO.o_iRequestPLCPC:=2;
		ELSE
			CommunicationIO.o_iRequestPLCPC:=1;
		END_IF;
ELSE
		IF ConveyorIO.xEmpty AND CommunicationIO.i_xExtraCondition THEN
			CommunicationIO.o_iRequestPLCPC:=2;
		ELSE
			CommunicationIO.o_iRequestPLCPC:=1;
		END_IF;
END_IF;	
(*出库段线体*)
(*//请求确认*)
CASE CommunicationIO.i_iResponsPCPLC OF 
	0:;
	1:;(*//复位*)
	2:(*//读码（入库申请）成功*)
	o_xReqSuccess:=1;
	3:(*//取放货完成*)
	ConveyorIO.xPutInto:=1; 
	4:(*//旋转*)
	o_xReqSuccess:=1;
	ConveyorIO.xPutInto:=1; 
	5:(*//不旋转*)
	o_xReqSuccess:=1;
	ConveyorIO.xPutInto:=1; 
	101:(*//条码空*)
	o_iErrorNub:=101;
	o_xError:=1;
	102:(*//条码规则检验失败*)
	o_iErrorNub:=102;
	o_xError:=1;
	103:(*//步号校验失败*)
	o_iErrorNub:=103;
	o_xError:=1;
	104:(*//无库位可用*)
	o_iErrorNub:=104;
	o_xError:=1;
	105:(*//路径选择失败*)
	o_iErrorNub:=105;
	o_xError:=1;
	106:(*//控制ID错误*)
	o_iErrorNub:=106;
	o_xError:=1;
	107:(*//叠盘计数不一致*)
	o_iErrorNub:=107;
	o_xError:=1;
END_CASE;
(*IF LDP(TRUE,CommunicationIO.i_iResponsPCPLC=3
			OR CommunicationIO.i_iResponsPCPLC =4
			OR CommunicationIO.i_iResponsPCPLC =5 ) THEN
	ConveyorIO.xPutInto:=1;
END_IF;*)
IF LDP(TRUE,CommunicationIO.i_iResponsPCPLC <> 3
			AND CommunicationIO.i_iResponsPCPLC <>4
			AND CommunicationIO.i_iResponsPCPLC <>5 ) THEN
	ConveyorIO.xPutInto:=0;
END_IF;
IF CommunicationIO.i_iResponsPCPLC <> 2 
	AND CommunicationIO.i_iResponsPCPLC <>4
	AND CommunicationIO.i_iResponsPCPLC <>5 THEN
	o_xReqSuccess:=0;
END_IF;
IF CommunicationIO.i_iResponsPCPLC < 100 THEN
	o_iErrorNub:=0;
	o_xError:=0;
END_IF;

(*//读写标志位写入数据*)
IF ConveyorIO.diDesConveyor<>ConveyorIO.diDeviceID THEN
	IF LDP(TRUE,CommunicationIO.i_iReadWriteFlagPCPLC = 1) THEN
		ConveyorIO.iTaskID := CommunicationIO.i_iTaskIDPCPLC;
		ConveyorIO.diDesConveyor := CommunicationIO.i_diDestinationDevicePCPLC;
		ConveyorIO.iProductCategory :=CommunicationIO.i_iProductIDPCPLC;
	END_IF;
END_IF;
(*//数据校验，并返回握手信号*)
IF CommunicationIO.i_iReadWriteFlagPCPLC = 1 
	AND ConveyorIO.iTaskID<>0
	AND ConveyorIO.diDesConveyor<>0 
	(*AND ConveyorIO.iProductCategory<>0 *)
	THEN
	CommunicationIO.o_iReadWriteFlagPLCPC:=2;
	(*处理标志位为2时，返回一个2*)
	ELSIF CommunicationIO.i_iTaskProcessFlagPCPLC=2 THEN
		CommunicationIO.o_iReadWriteFlagPLCPC:=2;
	ELSE
	CommunicationIO.o_iReadWriteFlagPLCPC:=1;
END_IF;

(*//数据校验*)
IF CommunicationIO.i_iReadWriteFlagPCPLC = 1 
	AND (ConveyorIO.iTaskID<>0
	OR ConveyorIO.diDesConveyor<>0 )
	(*OR ConveyorIO.iProductCategory<>0) *)
	THEN
	o_iErrorNub:=50;(*//任务数据不完整*)
END_IF;
(*//设备状态*)
IF ConveyorIO.diDesConveyor = ConveyorIO.diDeviceID 
		AND (ldp(TRUE,NOT ConveyorIO.xEmpty AND CommunicationIO.i_xExtraCondition) 
		OR (g_diDeviceIDSelect=ConveyorIO.diDeviceID AND g_xInsertTask))(*插入任务时，同时报一次完成*)
		THEN(*//目标地址=当前地址，表示是终点设备，有料就上传数据，报完成*)
	CommunicationIO.o_iDeviceStatusPLCPC:=3;(*//任务完成*)
	CommunicationIO.o_iProductIDPLCPC:=ConveyorIO.iProductCategory;(*//条码后四位上传*)
	CommunicationIO.o_iTaskIDPLCPC:=ConveyorIO.iTaskID;(*//任务号上传*)
	CommunicationIO.o_iRequestPLCPC:=2;(*发送入库请求*)
ELSIF ConveyorIO.diDesConveyor = ConveyorIO.diDeviceID AND LDp(TRUE,CommunicationIO.i_iTaskProcessFlagPCPLC=1)	
	THEN	(*//目标地址=当前地址，表示是终点设备，上位机给完成信号，就复位信号*)
	CommunicationIO.o_iDeviceStatusPLCPC:=1;
	CommunicationIO.o_iProductIDPLCPC:=0;(*//条码号复位*)
		CommunicationIO.o_iTaskIDPLCPC:=0;(*//任务号复位*)
ELSIF 	ConveyorIO.diDesConveyor <>ConveyorIO.diDeviceID AND ConveyorIO.xEmpty THEN(*非终点设备，无料就复位*)
	CommunicationIO.o_iDeviceStatusPLCPC:=1;
ELSIF ConveyorIO.xBusy THEN
	CommunicationIO.o_iDeviceStatusPLCPC:=2;(*//工作中*)
ELSIF ConveyorIO.xError THEN
	CommunicationIO.o_iDeviceStatusPLCPC:=4;(*//故障*)	
END_IF;
IF NOT g_xAuto THEN
	CommunicationIO.o_iDeviceStatusPLCPC:=0;
	CommunicationIO.o_iEmptyPLCPC:=0;
	CommunicationIO.o_iFolderNumberPLCPC:=0;
	CommunicationIO.o_iForceInportPLCPC:=0;
	CommunicationIO.o_iProductIDPLCPC:=0;
	CommunicationIO.o_iReadWriteFlagPLCPC:=0;
	CommunicationIO.o_iRequestPLCPC:=0;
	CommunicationIO.o_iTaskIDPLCPC:=0;
END_IF;
END_FUNCTION_BLOCK

FUNCTION_BLOCK ConveyorOld
VAR
  m_xPresentDelay : BOOL;  (* 有无判断延时 *)
  m_xLoadDelayOut : BOOL;  (* 上料延时输出 *)
  m_xInitial : BOOL;  (* 初始化 *)
  m_tUnloadTimer : TIME;  (* 下料计时器 *)
  m_tPresentDelayCurrentTime : TIME;
  m_tonUnloadAlam : TON;  (* 下料报警定时器 *)
  m_tonPresentDelay : TON;  (* 物料有无判断延时，防止误动作 *)
  m_tonNotArriveAlarm : TON;  (* 未到达报警计时 *)
  m_tonLoadDelay : TON;  (* 上料延时 *)
  m_tNotArriveCurrentTime : TIME;  (* 未到达报警计时当前时间 *)
  m_tLoadTimer : TIME;  (* 上料计时器 *)
  iStep : INT;  (* 上料步骤 *)
  m_wStateWord : INT;
END_VAR
VAR_IN_OUT
  ConveyorMotor : ConveyorIO;  (* 输送线输入输出 *)
END_VAR
VAR
  m_tonZoneClear : TON;  (* 初始化清除 *)
  m_tZoneClearCurrentTime : TIME;  (* 初始化清除当前时间 *)
  m_xAutoClear : BOOL;  (* 初始化清除标志位 *)
  m_xZoneClearDone : BOOL;  (* 初始化清除完成 *)
END_VAR
(*////////////////////////////////////////////////////////////////////////////////////////////////////////////
//传输线控制FB块，可控制单方向线体，双向旋转线体，支持双向上下料            
//线体初始化后为空的情况下输入xLoad信号即可进行上料动作，使用xLoadCCW信号可反方向上料
//增加了产品信息和产品种类的储存，当传输线为空和上料进行标志位为零的情况下清除产品信息和产品种类
//使用方式是在置位xLoad信号后，把产品信息和产品种类传入，等下料后自动清零
//线体不为空的情况下使用xUnload信号可进行下料动作，物料有无传感器的下降沿后出发计时器，延时断开传输线旋转
//单方向传输线体把xLoadCCW、xUnloadCCW设置为零，双向线体上料方向和下料反向的,方向固定的 把xUnloadCCW设置为1
//双方向线体双向都能上下料的要根据上料的方向来设置xLoadCCW,xUnloadCCW
//增加工作中信号xBusy当电机正转 显示为工作中
//增加上下料超时报警，xLoadAlarm，xUnloadAlarm，设定时间在LOAD_UNLOAD_TIME常量上，现在设置的为30秒
//增加xPutInto信号，用于直接投入的物料，检测开关感应到后，直接进入下料流程，上升沿有效
//离开延时改为变量 iLeaveDelay 默认为0 离开检测开关离输送线尾端比较远的线体需要根据情况设定100ms为单位
//增加初始化标志位，增加进入延时时间，初始化为进入延时时间为0 ，离开延时时间为2S，通过外围接口可以更改
//修改信息  修改后请增加版本
//12-17进行了优化，增加了未到达报警，当物料未传送到下一设备，就报未到达报警，使用xNextRun标志位制作，没有正常到达
//第0步，不能跳转到第一步把标志位复位，即出现中断情况，2秒后报警
//修改信息  修改后请增加版本
上料延时增加为50ms防止干扰信号
nextrun信号在 第三步也要复位
增加限位报警
增加超宽报警
增加产品型号输出在下料的时候把产品型号输送给下一段线体
增加线体单独复位
增加任务插入功能配合全局变量
增加暂停功能
增加线体状态字显示  0 空闲 1：有料  2 工作中  3  超限报警 4 超宽报警  5 未到达报警  6 下料超时报警
空料判断放在自动前，进行有无报警判断，然后跳转
修改超限报警，与尺寸检测报警
初始化清除线体标志位xZoneClear
ZPA zero pressure accumulation  Term that describes the Conveyor controls and mechanical scheme that will 
cause loads to queue on a conveyor in discrete zones such that loads do not touch each other(wrapped boxed tray tote carton)
//YAO      V1.0
///////////////////////////////////////////////////////////////////////////////////////////////////////////
(*********************************************************)
(*//初始化，
//上料延时位0S，下料报警延时为30S
//下料延时设一个比较大的时间，主要依靠xunload标志位来停止输送线，特殊情况可以用延时来停止物流线下料
//设置时间大的时候计时器会失效*)